// TIA Portal project "Tes simulation extract_V15.1" (V15.1) (continued)
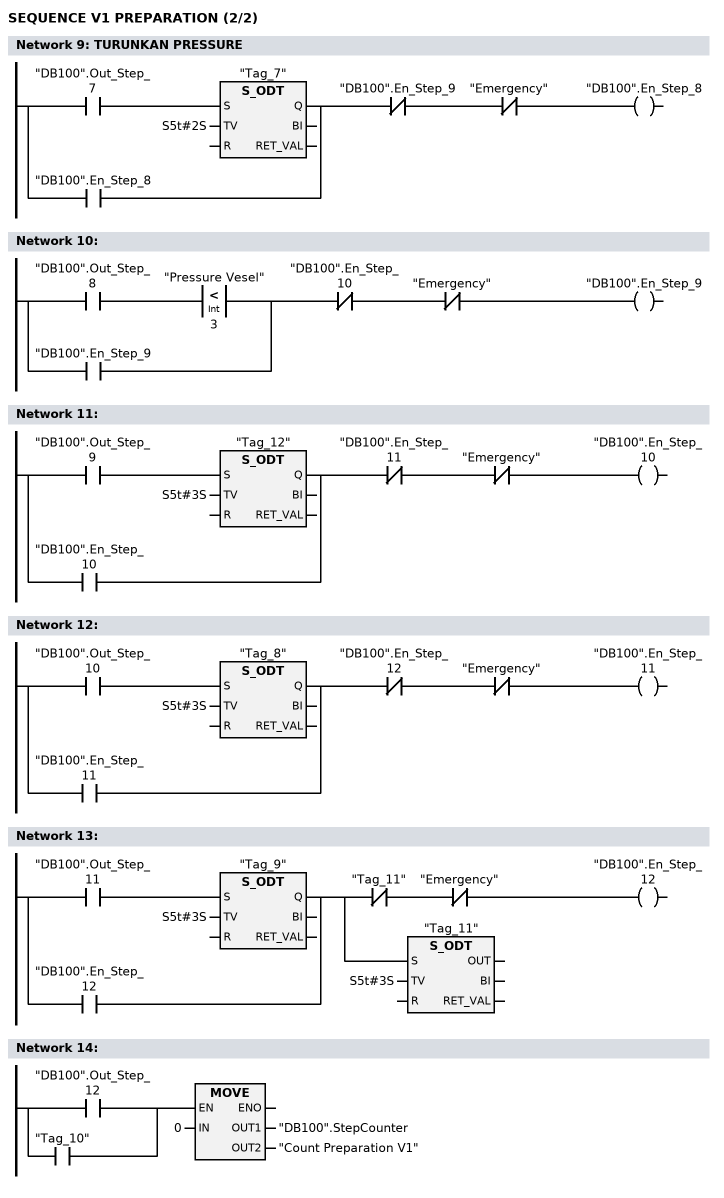
   RUNG wire#powerrail
      Contact( "DB100".Out_Step_7 )
      S_ODT(T_NO := "Tag_7", TV := S5t#2S, R :=, BI =>, RET_VAL =>)
      wire#w1
      I_Contact( "DB100".En_Step_9 )
      I_Contact( "Emergency" )
      Coil( "DB100".En_Step_8 )
   END_RUNG
   RUNG wire#powerrail
      Contact( "DB100".En_Step_8 )
   END_RUNG wire#w1
   // the same network as SCL:
   #_s5time1 := S_ODT(T_NO := "Tag_7", S := "DB100".Out_Step_7, TV := S5t#2S, Q => #_w1);
   "DB100".En_Step_8 := (#_w1 OR "DB100".En_Step_8) AND NOT "DB100".En_Step_9 AND NOT "Emergency";
END_REGION

REGION Network 10
   RUNG wire#powerrail
      Contact( "DB100".Out_Step_8 )
      { S7_Templates := "SrcType := Int" } LT_Contact(in1 := "Pressure Vesel", in2 := 3)
      wire#w1
      I_Contact( "DB100".En_Step_10 )
      I_Contact( "Emergency" )
      Coil( "DB100".En_Step_9 )
   END_RUNG
   RUNG wire#powerrail
      Contact( "DB100".En_Step_9 )
   END_RUNG wire#w1
   // the same network as SCL:
   "DB100".En_Step_9 := (("DB100".Out_Step_8 AND ("Pressure Vesel" < 3)) OR "DB100".En_Step_9) AND NOT "DB100".En_Step_10 AND NOT "Emergency";
END_REGION

REGION Network 11
   RUNG wire#powerrail
      Contact( "DB100".Out_Step_9 )
      S_ODT(T_NO := "Tag_12", TV := S5t#3S, R :=, BI =>, RET_VAL =>)
      wire#w1
      I_Contact( "DB100".En_Step_11 )
      I_Contact( "Emergency" )
      Coil( "DB100".En_Step_10 )
   END_RUNG
   RUNG wire#powerrail
      Contact( "DB100".En_Step_10 )
   END_RUNG wire#w1
   // the same network as SCL:
   #_s5time1 := S_ODT(T_NO := "Tag_12", S := "DB100".Out_Step_9, TV := S5t#3S, Q => #_w1);
   "DB100".En_Step_10 := (#_w1 OR "DB100".En_Step_10) AND NOT "DB100".En_Step_11 AND NOT "Emergency";
END_REGION

REGION Network 12
   RUNG wire#powerrail
      Contact( "DB100".Out_Step_10 )
      S_ODT(T_NO := "Tag_8", TV := S5t#3S, R :=, BI =>, RET_VAL =>)
      wire#w1
      I_Contact( "DB100".En_Step_12 )
      I_Contact( "Emergency" )
      Coil( "DB100".En_Step_11 )
   END_RUNG
   RUNG wire#powerrail
      Contact( "DB100".En_Step_11 )
   END_RUNG wire#w1
   // the same network as SCL:
   #_s5time1 := S_ODT(T_NO := "Tag_8", S := "DB100".Out_Step_10, TV := S5t#3S, Q => #_w1);
   "DB100".En_Step_11 := (#_w1 OR "DB100".En_Step_11) AND NOT "DB100".En_Step_12 AND NOT "Emergency";
END_REGION

REGION Network 13
   RUNG wire#powerrail
      Contact( "DB100".Out_Step_11 )
      S_ODT(T_NO := "Tag_9", TV := S5t#3S, R :=, BI =>, RET_VAL =>)
      wire#w1
      I_Contact( "Tag_11" )
      I_Contact( "Emergency" )
      Coil( "DB100".En_Step_12 )
   END_RUNG
   RUNG wire#powerrail
      Contact( "DB100".En_Step_12 )
   END_RUNG wire#w1
   RUNG wire#w1
      S_ODT(T_NO := "Tag_11", TV := S5t#3S, R :=, BI =>, RET_VAL =>)
   END_RUNG
   // the same network as SCL:
   #_s5time1 := S_ODT(T_NO := "Tag_9", S := "DB100".Out_Step_11, TV := S5t#3S, Q => #_w1);
   #_w2 := #_w1 OR "DB100".En_Step_12;
   "DB100".En_Step_12 := #_w2 AND NOT "Tag_11" AND NOT "Emergency";
   #_s5time2 := S_ODT(T_NO := "Tag_11", S := #_w2, TV := S5t#3S);
END_REGION

REGION Network 14
   RUNG wire#powerrail
      Contact( "DB100".Out_Step_12 )
      wire#w1
      Move(in := 0, out1 => "DB100".StepCounter, out2 => "Count Preparation V1")
   END_RUNG
   RUNG wire#powerrail
      Contact( "Tag_10" )
   END_RUNG wire#w1
   // the same network as SCL:
   IF "DB100".Out_Step_12 OR "Tag_10" THEN
       "DB100".StepCounter := 0;
       "Count Preparation V1" := 0;
   END_IF;
END_REGION
END_FUNCTION

FUNCTION "VESSEL 1 PREPARATION" : Void   // FC2, LAD
{ S7_Optimized_Access := 'TRUE' }
VERSION : 0.1
   VAR_TEMP   // added for the SCL form of the ladder/FBD networks
      _w1 : Bool;
      _w2 : Bool;
      _w3 : Bool;
      _w4 : Bool;
   END_VAR
BEGIN

REGION Network 1: NAIKAN PRESSURE STEAM
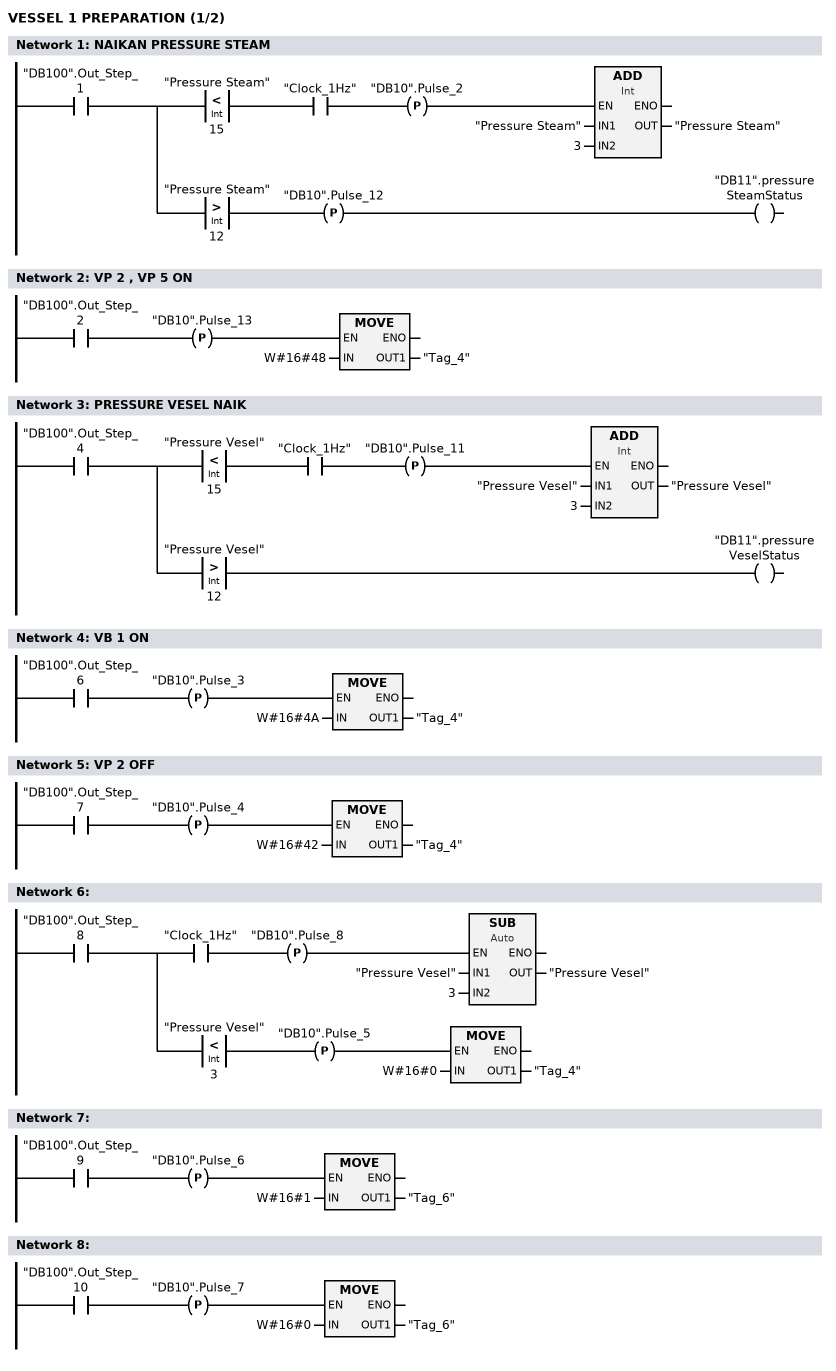
   RUNG wire#powerrail
      Contact( "DB100".Out_Step_1 )
      wire#w1
      { S7_Templates := "SrcType := Int" } LT_Contact(in1 := "Pressure Steam", in2 := 15)
      Contact( "Clock_1Hz" )
      P_Trig( "DB10".Pulse_2 )
      { S7_Templates := "SrcType := Int" } Add(in1 := "Pressure Steam", in2 := 3, out => "Pressure Steam")
   END_RUNG
   RUNG wire#w1
      { S7_Templates := "SrcType := Int" } GT_Contact(in1 := "Pressure Steam", in2 := 12)
      P_Trig( "DB10".Pulse_12 )
      Coil( "DB11".pressureSteamStatus )
   END_RUNG
   // the same network as SCL:
   #_w1 := "DB100".Out_Step_1 AND ("Pressure Steam" < 15) AND "Clock_1Hz";
   #_w2 := #_w1 AND NOT "DB10".Pulse_2;   // rising edge
   "DB10".Pulse_2 := #_w1;
   IF #_w2 THEN "Pressure Steam" := "Pressure Steam" + 3; END_IF;
   #_w3 := "DB100".Out_Step_1 AND ("Pressure Steam" > 12);
   #_w4 := #_w3 AND NOT "DB10".Pulse_12;   // rising edge
   "DB10".Pulse_12 := #_w3;
   "DB11".pressureSteamStatus := #_w4;
END_REGION

REGION Network 2: VP 2 , VP 5 ON
   RUNG wire#powerrail
      Contact( "DB100".Out_Step_2 )
      P_Trig( "DB10".Pulse_13 )
      Move(in := W#16#48, out1 => "Tag_4")
   END_RUNG
   // the same network as SCL:
   #_w1 := "DB100".Out_Step_2 AND NOT "DB10".Pulse_13;   // rising edge
   "DB10".Pulse_13 := "DB100".Out_Step_2;
   IF #_w1 THEN "Tag_4" := W#16#48; END_IF;
END_REGION

REGION Network 3: PRESSURE VESEL NAIK
   RUNG wire#powerrail
      Contact( "DB100".Out_Step_4 )
      wire#w1
      { S7_Templates := "SrcType := Int" } LT_Contact(in1 := "Pressure Vesel", in2 := 15)
      Contact( "Clock_1Hz" )
      P_Trig( "DB10".Pulse_11 )
      { S7_Templates := "SrcType := Int" } Add(in1 := "Pressure Vesel", in2 := 3, out => "Pressure Vesel")
   END_RUNG
   RUNG wire#w1
      { S7_Templates := "SrcType := Int" } GT_Contact(in1 := "Pressure Vesel", in2 := 12)
      Coil( "DB11".pressureVeselStatus )
   END_RUNG
   // the same network as SCL:
   #_w1 := "DB100".Out_Step_4 AND ("Pressure Vesel" < 15) AND "Clock_1Hz";
   #_w2 := #_w1 AND NOT "DB10".Pulse_11;   // rising edge
   "DB10".Pulse_11 := #_w1;
   IF #_w2 THEN "Pressure Vesel" := "Pressure Vesel" + 3; END_IF;
   "DB11".pressureVeselStatus := "DB100".Out_Step_4 AND ("Pressure Vesel" > 12);
END_REGION

REGION Network 4: VB 1 ON
   RUNG wire#powerrail
      Contact( "DB100".Out_Step_6 )
      P_Trig( "DB10".Pulse_3 )
      Move(in := W#16#4A, out1 => "Tag_4")
   END_RUNG
   // the same network as SCL:
   #_w1 := "DB100".Out_Step_6 AND NOT "DB10".Pulse_3;   // rising edge
   "DB10".Pulse_3 := "DB100".Out_Step_6;
   IF #_w1 THEN "Tag_4" := W#16#4A; END_IF;
END_REGION

REGION Network 5: VP 2 OFF
   RUNG wire#powerrail
      Contact( "DB100".Out_Step_7 )
      P_Trig( "DB10".Pulse_4 )
      Move(in := W#16#42, out1 => "Tag_4")
   END_RUNG
   // the same network as SCL:
   #_w1 := "DB100".Out_Step_7 AND NOT "DB10".Pulse_4;   // rising edge
   "DB10".Pulse_4 := "DB100".Out_Step_7;
   IF #_w1 THEN "Tag_4" := W#16#42; END_IF;
END_REGION

REGION Network 6
   RUNG wire#powerrail
      Contact( "DB100".Out_Step_8 )
      wire#w1
      Contact( "Clock_1Hz" )
      P_Trig( "DB10".Pulse_8 )
      Sub(in1 := "Pressure Vesel", in2 := 3, out => "Pressure Vesel")
   END_RUNG
   RUNG wire#w1
      { S7_Templates := "SrcType := Int" } LT_Contact(in1 := "Pressure Vesel", in2 := 3)
      P_Trig( "DB10".Pulse_5 )
      Move(in := W#16#0, out1 => "Tag_4")
   END_RUNG
   // the same network as SCL:
   #_w1 := "DB100".Out_Step_8 AND "Clock_1Hz";
   #_w2 := #_w1 AND NOT "DB10".Pulse_8;   // rising edge
   "DB10".Pulse_8 := #_w1;
   IF #_w2 THEN "Pressure Vesel" := "Pressure Vesel" - 3; END_IF;
   #_w3 := "DB100".Out_Step_8 AND ("Pressure Vesel" < 3);
   #_w4 := #_w3 AND NOT "DB10".Pulse_5;   // rising edge
   "DB10".Pulse_5 := #_w3;
   IF #_w4 THEN "Tag_4" := W#16#0; END_IF;
END_REGION

REGION Network 7
   RUNG wire#powerrail
      Contact( "DB100".Out_Step_9 )
      P_Trig( "DB10".Pulse_6 )
      Move(in := W#16#1, out1 => "Tag_6")
   END_RUNG
   // the same network as SCL:
   #_w1 := "DB100".Out_Step_9 AND NOT "DB10".Pulse_6;   // rising edge
   "DB10".Pulse_6 := "DB100".Out_Step_9;
   IF #_w1 THEN "Tag_6" := W#16#1; END_IF;
END_REGION

REGION Network 8
   RUNG wire#powerrail
      Contact( "DB100".Out_Step_10 )
      P_Trig( "DB10".Pulse_7 )
      Move(in := W#16#0, out1 => "Tag_6")
   END_RUNG
   // the same network as SCL:
   #_w1 := "DB100".Out_Step_10 AND NOT "DB10".Pulse_7;   // rising edge
   "DB10".Pulse_7 := "DB100".Out_Step_10;
   IF #_w1 THEN "Tag_6" := W#16#0; END_IF;
END_REGION

REGION Network 9
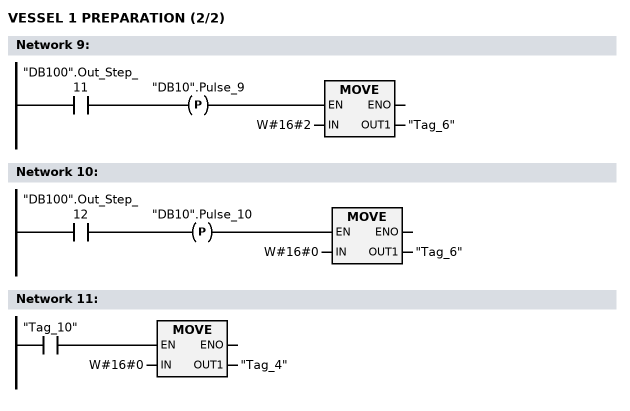
   RUNG wire#powerrail
      Contact( "DB100".Out_Step_11 )
      P_Trig( "DB10".Pulse_9 )
      Move(in := W#16#2, out1 => "Tag_6")
   END_RUNG
   // the same network as SCL:
   #_w1 := "DB100".Out_Step_11 AND NOT "DB10".Pulse_9;   // rising edge
   "DB10".Pulse_9 := "DB100".Out_Step_11;
   IF #_w1 THEN "Tag_6" := W#16#2; END_IF;
END_REGION

REGION Network 10
   RUNG wire#powerrail
      Contact( "DB100".Out_Step_12 )
      P_Trig( "DB10".Pulse_10 )
      Move(in := W#16#0, out1 => "Tag_6")
   END_RUNG
   // the same network as SCL:
   #_w1 := "DB100".Out_Step_12 AND NOT "DB10".Pulse_10;   // rising edge
   "DB10".Pulse_10 := "DB100".Out_Step_12;
   IF #_w1 THEN "Tag_6" := W#16#0; END_IF;
END_REGION

REGION Network 11
   RUNG wire#powerrail
      Contact( "Tag_10" )
      Move(in := W#16#0, out1 => "Tag_4")
   END_RUNG
   // the same network as SCL:
   IF "Tag_10" THEN "Tag_4" := W#16#0; END_IF;
END_REGION
END_FUNCTION

FUNCTION "ISI VESEL" : Void   // FC3, LAD
{ S7_Optimized_Access := 'TRUE' }
VERSION : 0.1
   VAR_TEMP   // added for the SCL form of the ladder/FBD networks
      _w1 : Bool;
      _w2 : Bool;
      _s5time1 : S5Time;
   END_VAR
BEGIN

REGION Network 1: ISI VESEL 1
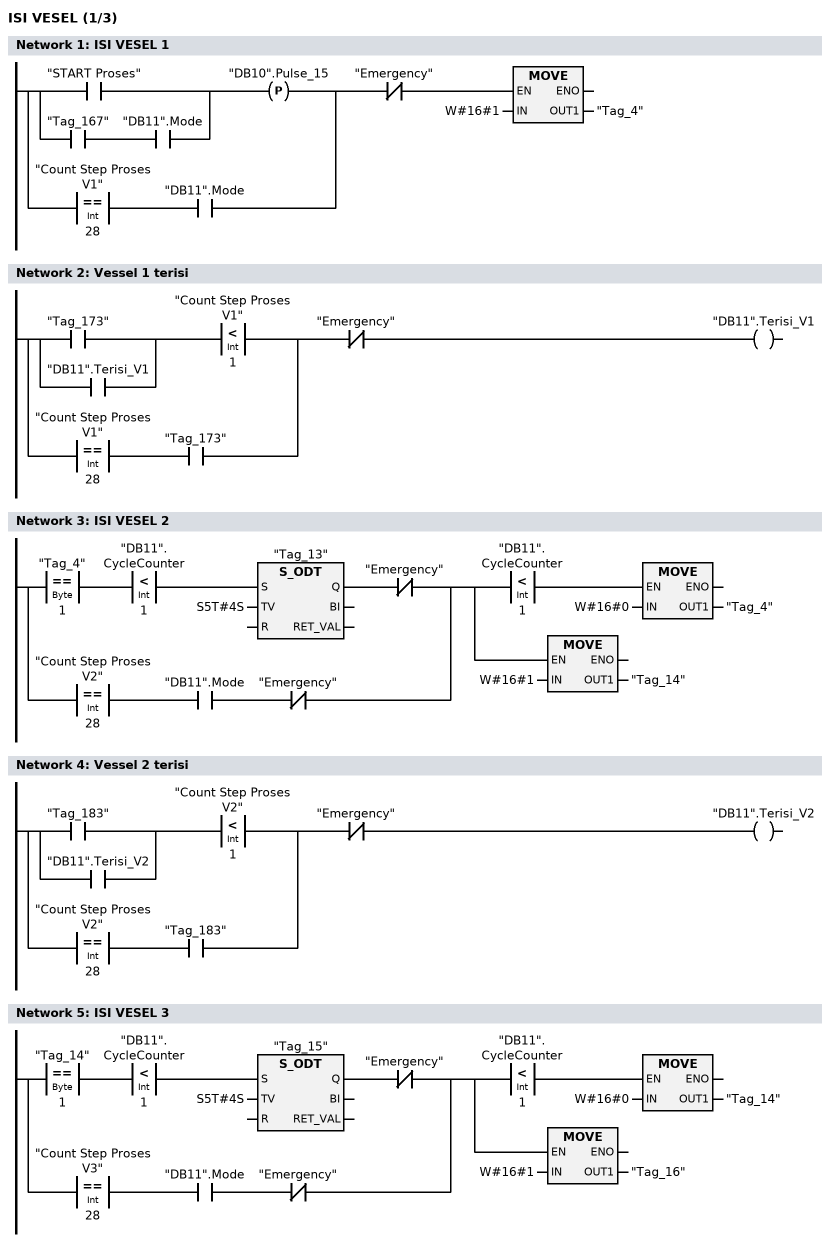
   RUNG wire#powerrail
      Contact( "START Proses" )
      wire#w1
      P_Trig( "DB10".Pulse_15 )
      wire#w2
      I_Contact( "Emergency" )
      Move(in := W#16#1, out1 => "Tag_4")
   END_RUNG
   RUNG wire#powerrail
      Contact( "Tag_167" )
      Contact( "DB11".Mode )
   END_RUNG wire#w1
   RUNG wire#powerrail
      { S7_Templates := "SrcType := Int" } EQ_Contact(in1 := "Count Step Proses V1", in2 := 28)
      Contact( "DB11".Mode )
   END_RUNG wire#w2
   // the same network as SCL:
   #_w1 := "START Proses" OR ("Tag_167" AND "DB11".Mode);
   #_w2 := #_w1 AND NOT "DB10".Pulse_15;   // rising edge
   "DB10".Pulse_15 := #_w1;
   IF (#_w2 OR (("Count Step Proses V1" = 28) AND "DB11".Mode)) AND NOT "Emergency" THEN
       "Tag_4" := W#16#1;
   END_IF;
END_REGION

REGION Network 2: Vessel 1 terisi
   RUNG wire#powerrail
      Contact( "Tag_173" )
      wire#w1
      { S7_Templates := "SrcType := Int" } LT_Contact(in1 := "Count Step Proses V1", in2 := 1)
      wire#w2
      I_Contact( "Emergency" )
      Coil( "DB11".Terisi_V1 )
   END_RUNG
   RUNG wire#powerrail
      Contact( "DB11".Terisi_V1 )
   END_RUNG wire#w1
   RUNG wire#powerrail
      { S7_Templates := "SrcType := Int" } EQ_Contact(in1 := "Count Step Proses V1", in2 := 28)
      Contact( "Tag_173" )
   END_RUNG wire#w2
   // the same network as SCL:
   "DB11".Terisi_V1 := ((("Tag_173" OR "DB11".Terisi_V1) AND ("Count Step Proses V1" < 1)) OR (("Count Step Proses V1" = 28) AND "Tag_173")) AND NOT "Emergency";
END_REGION

REGION Network 3: ISI VESEL 2
   RUNG wire#powerrail
      { S7_Templates := "SrcType := Byte" } EQ_Contact(in1 := "Tag_4", in2 := 1)
      { S7_Templates := "SrcType := Int" } LT_Contact(in1 := "DB11".CycleCounter, in2 := 1)
      S_ODT(T_NO := "Tag_13", TV := S5T#4S, R :=, BI =>, RET_VAL =>)
      I_Contact( "Emergency" )
      wire#w1
      { S7_Templates := "SrcType := Int" } LT_Contact(in1 := "DB11".CycleCounter, in2 := 1)
      Move(in := W#16#0, out1 => "Tag_4")
   END_RUNG
   RUNG wire#powerrail
      { S7_Templates := "SrcType := Int" } EQ_Contact(in1 := "Count Step Proses V2", in2 := 28)
      Contact( "DB11".Mode )
      I_Contact( "Emergency" )
   END_RUNG wire#w1
   RUNG wire#w1
      Move(in := W#16#1, out1 => "Tag_14")
   END_RUNG
   // the same network as SCL:
   #_s5time1 := S_ODT(T_NO := "Tag_13",
                      S := ("Tag_4" = 1) AND ("DB11".CycleCounter < 1),
                      TV := S5T#4S,
                      Q => #_w1);
   #_w2 := (#_w1 AND NOT "Emergency") OR (("Count Step Proses V2" = 28) AND "DB11".Mode AND NOT "Emergency");
   IF #_w2 AND ("DB11".CycleCounter < 1) THEN "Tag_4" := W#16#0; END_IF;
   IF #_w2 THEN "Tag_14" := W#16#1; END_IF;
END_REGION

REGION Network 4: Vessel 2 terisi
   RUNG wire#powerrail
      Contact( "Tag_183" )
      wire#w1
      { S7_Templates := "SrcType := Int" } LT_Contact(in1 := "Count Step Proses V2", in2 := 1)
      wire#w2
      I_Contact( "Emergency" )
      Coil( "DB11".Terisi_V2 )
   END_RUNG
   RUNG wire#powerrail
      Contact( "DB11".Terisi_V2 )
   END_RUNG wire#w1
   RUNG wire#powerrail
      { S7_Templates := "SrcType := Int" } EQ_Contact(in1 := "Count Step Proses V2", in2 := 28)
      Contact( "Tag_183" )
   END_RUNG wire#w2
   // the same network as SCL:
   "DB11".Terisi_V2 := ((("Tag_183" OR "DB11".Terisi_V2) AND ("Count Step Proses V2" < 1)) OR (("Count Step Proses V2" = 28) AND "Tag_183")) AND NOT "Emergency";
END_REGION

REGION Network 5: ISI VESEL 3
   RUNG wire#powerrail
      { S7_Templates := "SrcType := Byte" } EQ_Contact(in1 := "Tag_14", in2 := 1)
      { S7_Templates := "SrcType := Int" } LT_Contact(in1 := "DB11".CycleCounter, in2 := 1)
      S_ODT(T_NO := "Tag_15", TV := S5T#4S, R :=, BI =>, RET_VAL =>)
      I_Contact( "Emergency" )
      wire#w1
      { S7_Templates := "SrcType := Int" } LT_Contact(in1 := "DB11".CycleCounter, in2 := 1)
      Move(in := W#16#0, out1 => "Tag_14")
   END_RUNG
   RUNG wire#powerrail
      { S7_Templates := "SrcType := Int" } EQ_Contact(in1 := "Count Step Proses V3", in2 := 28)
      Contact( "DB11".Mode )
      I_Contact( "Emergency" )
   END_RUNG wire#w1
   RUNG wire#w1
      Move(in := W#16#1, out1 => "Tag_16")
   END_RUNG
   // the same network as SCL:
   #_s5time1 := S_ODT(T_NO := "Tag_15",
                      S := ("Tag_14" = 1) AND ("DB11".CycleCounter < 1),
                      TV := S5T#4S,
                      Q => #_w1);
   #_w2 := (#_w1 AND NOT "Emergency") OR (("Count Step Proses V3" = 28) AND "DB11".Mode AND NOT "Emergency");
   IF #_w2 AND ("DB11".CycleCounter < 1) THEN "Tag_14" := W#16#0; END_IF;
   IF #_w2 THEN "Tag_16" := W#16#1; END_IF;
END_REGION

REGION Network 6: Vessel 3 terisi
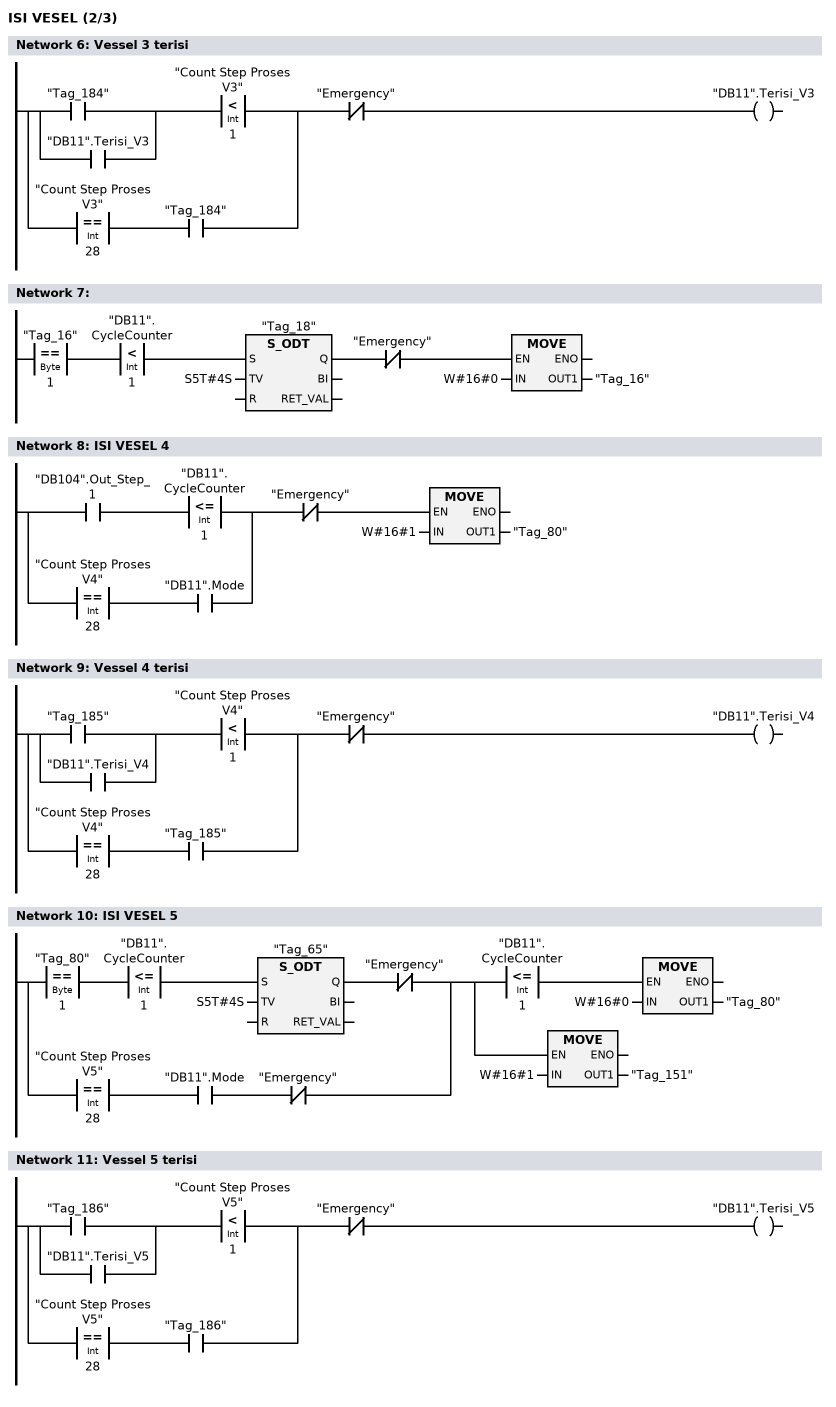
   RUNG wire#powerrail
      Contact( "Tag_184" )
      wire#w1
      { S7_Templates := "SrcType := Int" } LT_Contact(in1 := "Count Step Proses V3", in2 := 1)
      wire#w2
      I_Contact( "Emergency" )
      Coil( "DB11".Terisi_V3 )
   END_RUNG
   RUNG wire#powerrail
      Contact( "DB11".Terisi_V3 )
   END_RUNG wire#w1
   RUNG wire#powerrail
      { S7_Templates := "SrcType := Int" } EQ_Contact(in1 := "Count Step Proses V3", in2 := 28)
      Contact( "Tag_184" )
   END_RUNG wire#w2
   // the same network as SCL:
   "DB11".Terisi_V3 := ((("Tag_184" OR "DB11".Terisi_V3) AND ("Count Step Proses V3" < 1)) OR (("Count Step Proses V3" = 28) AND "Tag_184")) AND NOT "Emergency";
END_REGION

REGION Network 7
   RUNG wire#powerrail
      { S7_Templates := "SrcType := Byte" } EQ_Contact(in1 := "Tag_16", in2 := 1)
      { S7_Templates := "SrcType := Int" } LT_Contact(in1 := "DB11".CycleCounter, in2 := 1)
      S_ODT(T_NO := "Tag_18", TV := S5T#4S, R :=, BI =>, RET_VAL =>)
      I_Contact( "Emergency" )
      Move(in := W#16#0, out1 => "Tag_16")
   END_RUNG
   // the same network as SCL:
   #_s5time1 := S_ODT(T_NO := "Tag_18",
                      S := ("Tag_16" = 1) AND ("DB11".CycleCounter < 1),
                      TV := S5T#4S,
                      Q => #_w1);
   IF #_w1 AND NOT "Emergency" THEN "Tag_16" := W#16#0; END_IF;
END_REGION

REGION Network 8: ISI VESEL 4
   RUNG wire#powerrail
      Contact( "DB104".Out_Step_1 )
      { S7_Templates := "SrcType := Int" } LE_Contact(in1 := "DB11".CycleCounter, in2 := 1)
      wire#w1
      I_Contact( "Emergency" )
      Move(in := W#16#1, out1 => "Tag_80")
   END_RUNG
   RUNG wire#powerrail
      { S7_Templates := "SrcType := Int" } EQ_Contact(in1 := "Count Step Proses V4", in2 := 28)
      Contact( "DB11".Mode )
   END_RUNG wire#w1
   // the same network as SCL:
   IF (("DB104".Out_Step_1 AND ("DB11".CycleCounter <= 1)) OR (("Count Step Proses V4" = 28) AND "DB11".Mode)) AND NOT "Emergency" THEN
       "Tag_80" := W#16#1;
   END_IF;
END_REGION

REGION Network 9: Vessel 4 terisi
   RUNG wire#powerrail
      Contact( "Tag_185" )
      wire#w1
      { S7_Templates := "SrcType := Int" } LT_Contact(in1 := "Count Step Proses V4", in2 := 1)
      wire#w2
      I_Contact( "Emergency" )
      Coil( "DB11".Terisi_V4 )
   END_RUNG
   RUNG wire#powerrail
      Contact( "DB11".Terisi_V4 )
   END_RUNG wire#w1
   RUNG wire#powerrail
      { S7_Templates := "SrcType := Int" } EQ_Contact(in1 := "Count Step Proses V4", in2 := 28)
      Contact( "Tag_185" )
   END_RUNG wire#w2
   // the same network as SCL:
   "DB11".Terisi_V4 := ((("Tag_185" OR "DB11".Terisi_V4) AND ("Count Step Proses V4" < 1)) OR (("Count Step Proses V4" = 28) AND "Tag_185")) AND NOT "Emergency";
END_REGION

REGION Network 10: ISI VESEL 5
   RUNG wire#powerrail
      { S7_Templates := "SrcType := Byte" } EQ_Contact(in1 := "Tag_80", in2 := 1)
      { S7_Templates := "SrcType := Int" } LE_Contact(in1 := "DB11".CycleCounter, in2 := 1)
      S_ODT(T_NO := "Tag_65", TV := S5T#4S, R :=, BI =>, RET_VAL =>)
      I_Contact( "Emergency" )
      wire#w1
      { S7_Templates := "SrcType := Int" } LE_Contact(in1 := "DB11".CycleCounter, in2 := 1)
      Move(in := W#16#0, out1 => "Tag_80")
   END_RUNG
   RUNG wire#powerrail
      { S7_Templates := "SrcType := Int" } EQ_Contact(in1 := "Count Step Proses V5", in2 := 28)
      Contact( "DB11".Mode )
      I_Contact( "Emergency" )
   END_RUNG wire#w1
   RUNG wire#w1
      Move(in := W#16#1, out1 => "Tag_151")
   END_RUNG
   // the same network as SCL:
   #_s5time1 := S_ODT(T_NO := "Tag_65",
                      S := ("Tag_80" = 1) AND ("DB11".CycleCounter <= 1),
                      TV := S5T#4S,
                      Q => #_w1);
   #_w2 := (#_w1 AND NOT "Emergency") OR (("Count Step Proses V5" = 28) AND "DB11".Mode AND NOT "Emergency");
   IF #_w2 AND ("DB11".CycleCounter <= 1) THEN "Tag_80" := W#16#0; END_IF;
   IF #_w2 THEN "Tag_151" := W#16#1; END_IF;
END_REGION

REGION Network 11: Vessel 5 terisi
   RUNG wire#powerrail
      Contact( "Tag_186" )
      wire#w1
      { S7_Templates := "SrcType := Int" } LT_Contact(in1 := "Count Step Proses V5", in2 := 1)
      wire#w2
      I_Contact( "Emergency" )
      Coil( "DB11".Terisi_V5 )
   END_RUNG
   RUNG wire#powerrail
      Contact( "DB11".Terisi_V5 )
   END_RUNG wire#w1
   RUNG wire#powerrail
      { S7_Templates := "SrcType := Int" } EQ_Contact(in1 := "Count Step Proses V5", in2 := 28)
      Contact( "Tag_186" )
   END_RUNG wire#w2
   // the same network as SCL:
   "DB11".Terisi_V5 := ((("Tag_186" OR "DB11".Terisi_V5) AND ("Count Step Proses V5" < 1)) OR (("Count Step Proses V5" = 28) AND "Tag_186")) AND NOT "Emergency";
END_REGION

REGION Network 12: ISI VESEL 6
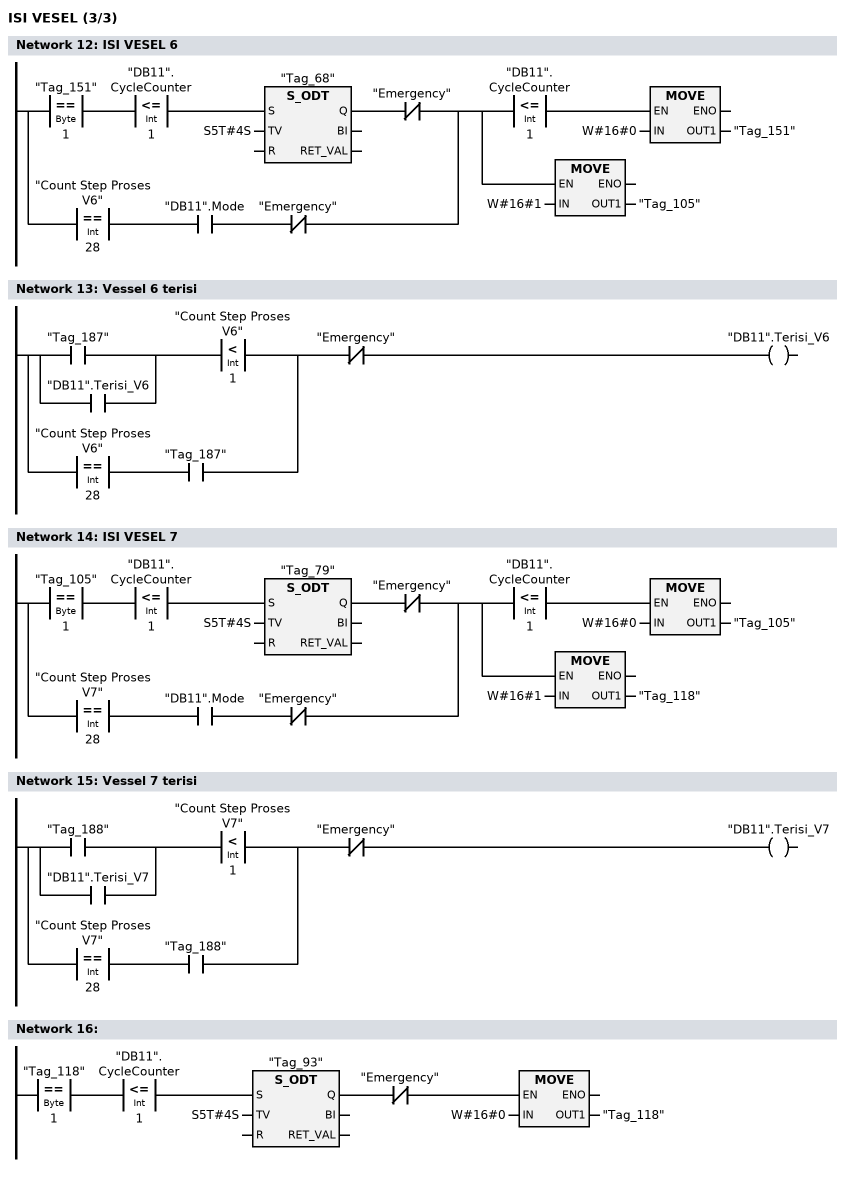
   RUNG wire#powerrail
      { S7_Templates := "SrcType := Byte" } EQ_Contact(in1 := "Tag_151", in2 := 1)
      { S7_Templates := "SrcType := Int" } LE_Contact(in1 := "DB11".CycleCounter, in2 := 1)
      S_ODT(T_NO := "Tag_68", TV := S5T#4S, R :=, BI =>, RET_VAL =>)
      I_Contact( "Emergency" )
      wire#w1
      { S7_Templates := "SrcType := Int" } LE_Contact(in1 := "DB11".CycleCounter, in2 := 1)
      Move(in := W#16#0, out1 => "Tag_151")
   END_RUNG
   RUNG wire#powerrail
      { S7_Templates := "SrcType := Int" } EQ_Contact(in1 := "Count Step Proses V6", in2 := 28)
      Contact( "DB11".Mode )
      I_Contact( "Emergency" )
   END_RUNG wire#w1
   RUNG wire#w1
      Move(in := W#16#1, out1 => "Tag_105")
   END_RUNG
   // the same network as SCL:
   #_s5time1 := S_ODT(T_NO := "Tag_68",
                      S := ("Tag_151" = 1) AND ("DB11".CycleCounter <= 1),
                      TV := S5T#4S,
                      Q => #_w1);
   #_w2 := (#_w1 AND NOT "Emergency") OR (("Count Step Proses V6" = 28) AND "DB11".Mode AND NOT "Emergency");
   IF #_w2 AND ("DB11".CycleCounter <= 1) THEN "Tag_151" := W#16#0; END_IF;
   IF #_w2 THEN "Tag_105" := W#16#1; END_IF;
END_REGION

REGION Network 13: Vessel 6 terisi
   RUNG wire#powerrail
      Contact( "Tag_187" )
      wire#w1
      { S7_Templates := "SrcType := Int" } LT_Contact(in1 := "Count Step Proses V6", in2 := 1)
      wire#w2
      I_Contact( "Emergency" )
      Coil( "DB11".Terisi_V6 )
   END_RUNG
   RUNG wire#powerrail
      Contact( "DB11".Terisi_V6 )
   END_RUNG wire#w1
   RUNG wire#powerrail
      { S7_Templates := "SrcType := Int" } EQ_Contact(in1 := "Count Step Proses V6", in2 := 28)
      Contact( "Tag_187" )
   END_RUNG wire#w2
   // the same network as SCL:
   "DB11".Terisi_V6 := ((("Tag_187" OR "DB11".Terisi_V6) AND ("Count Step Proses V6" < 1)) OR (("Count Step Proses V6" = 28) AND "Tag_187")) AND NOT "Emergency";
END_REGION

REGION Network 14: ISI VESEL 7
   RUNG wire#powerrail
      { S7_Templates := "SrcType := Byte" } EQ_Contact(in1 := "Tag_105", in2 := 1)
      { S7_Templates := "SrcType := Int" } LE_Contact(in1 := "DB11".CycleCounter, in2 := 1)
      S_ODT(T_NO := "Tag_79", TV := S5T#4S, R :=, BI =>, RET_VAL =>)
      I_Contact( "Emergency" )
      wire#w1
      { S7_Templates := "SrcType := Int" } LE_Contact(in1 := "DB11".CycleCounter, in2 := 1)
      Move(in := W#16#0, out1 => "Tag_105")
   END_RUNG
   RUNG wire#powerrail
      { S7_Templates := "SrcType := Int" } EQ_Contact(in1 := "Count Step Proses V7", in2 := 28)
      Contact( "DB11".Mode )
      I_Contact( "Emergency" )
   END_RUNG wire#w1
   RUNG wire#w1
      Move(in := W#16#1, out1 => "Tag_118")
   END_RUNG
   // the same network as SCL:
   #_s5time1 := S_ODT(T_NO := "Tag_79",
                      S := ("Tag_105" = 1) AND ("DB11".CycleCounter <= 1),
                      TV := S5T#4S,
                      Q => #_w1);
   #_w2 := (#_w1 AND NOT "Emergency") OR (("Count Step Proses V7" = 28) AND "DB11".Mode AND NOT "Emergency");
   IF #_w2 AND ("DB11".CycleCounter <= 1) THEN "Tag_105" := W#16#0; END_IF;
   IF #_w2 THEN "Tag_118" := W#16#1; END_IF;
END_REGION

REGION Network 15: Vessel 7 terisi
   RUNG wire#powerrail
      Contact( "Tag_188" )
      wire#w1
      { S7_Templates := "SrcType := Int" } LT_Contact(in1 := "Count Step Proses V7", in2 := 1)
      wire#w2
      I_Contact( "Emergency" )
      Coil( "DB11".Terisi_V7 )
   END_RUNG
   RUNG wire#powerrail
      Contact( "DB11".Terisi_V7 )
   END_RUNG wire#w1
   RUNG wire#powerrail
      { S7_Templates := "SrcType := Int" } EQ_Contact(in1 := "Count Step Proses V7", in2 := 28)
      Contact( "Tag_188" )
   END_RUNG wire#w2
   // the same network as SCL:
   "DB11".Terisi_V7 := ((("Tag_188" OR "DB11".Terisi_V7) AND ("Count Step Proses V7" < 1)) OR (("Count Step Proses V7" = 28) AND "Tag_188")) AND NOT "Emergency";
END_REGION

REGION Network 16
   RUNG wire#powerrail
      { S7_Templates := "SrcType := Byte" } EQ_Contact(in1 := "Tag_118", in2 := 1)
      { S7_Templates := "SrcType := Int" } LE_Contact(in1 := "DB11".CycleCounter, in2 := 1)
      S_ODT(T_NO := "Tag_93", TV := S5T#4S, R :=, BI =>, RET_VAL =>)
      I_Contact( "Emergency" )
      Move(in := W#16#0, out1 => "Tag_118")
   END_RUNG
   // the same network as SCL:
   #_s5time1 := S_ODT(T_NO := "Tag_93",
                      S := ("Tag_118" = 1) AND ("DB11".CycleCounter <= 1),
                      TV := S5T#4S,
                      Q => #_w1);
   IF #_w1 AND NOT "Emergency" THEN "Tag_118" := W#16#0; END_IF;
END_REGION
END_FUNCTION

FUNCTION "SUPPLY" : Void   // FC4, LAD
{ S7_Optimized_Access := 'TRUE' }
VERSION : 0.1
   VAR_TEMP   // added for the SCL form of the ladder/FBD networks
      _w1 : Bool;
      _w2 : Bool;
      _w3 : Bool;
      _w4 : Bool;
   END_VAR
BEGIN

REGION Network 1: BUKA CV AIR 1
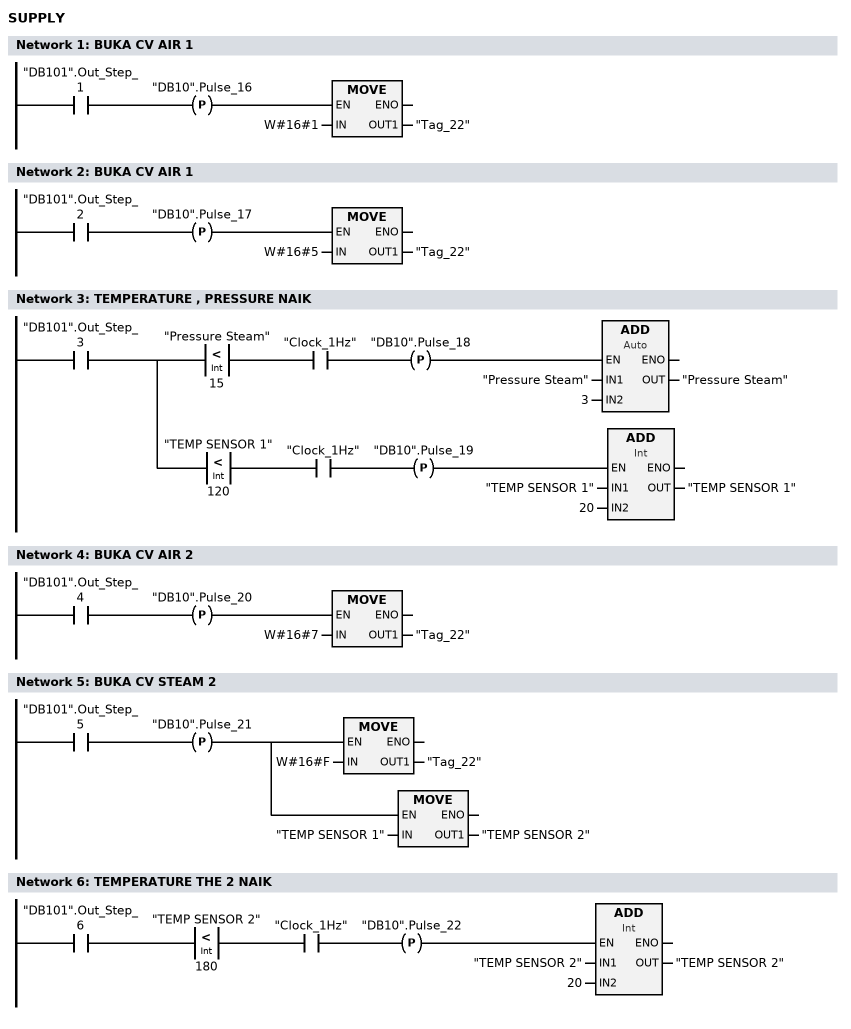
   RUNG wire#powerrail
      Contact( "DB101".Out_Step_1 )
      P_Trig( "DB10".Pulse_16 )
      Move(in := W#16#1, out1 => "Tag_22")
   END_RUNG
   // the same network as SCL:
   #_w1 := "DB101".Out_Step_1 AND NOT "DB10".Pulse_16;   // rising edge
   "DB10".Pulse_16 := "DB101".Out_Step_1;
   IF #_w1 THEN "Tag_22" := W#16#1; END_IF;
END_REGION

REGION Network 2: BUKA CV AIR 1
   RUNG wire#powerrail
      Contact( "DB101".Out_Step_2 )
      P_Trig( "DB10".Pulse_17 )
      Move(in := W#16#5, out1 => "Tag_22")
   END_RUNG
   // the same network as SCL:
   #_w1 := "DB101".Out_Step_2 AND NOT "DB10".Pulse_17;   // rising edge
   "DB10".Pulse_17 := "DB101".Out_Step_2;
   IF #_w1 THEN "Tag_22" := W#16#5; END_IF;
END_REGION

REGION Network 3: TEMPERATURE , PRESSURE NAIK
   RUNG wire#powerrail
      Contact( "DB101".Out_Step_3 )
      wire#w1
      { S7_Templates := "SrcType := Int" } LT_Contact(in1 := "Pressure Steam", in2 := 15)
      Contact( "Clock_1Hz" )
      P_Trig( "DB10".Pulse_18 )
      Add(in1 := "Pressure Steam", in2 := 3, out => "Pressure Steam")
   END_RUNG
   RUNG wire#w1
      { S7_Templates := "SrcType := Int" } LT_Contact(in1 := "TEMP SENSOR 1", in2 := 120)
      Contact( "Clock_1Hz" )
      P_Trig( "DB10".Pulse_19 )
      { S7_Templates := "SrcType := Int" } Add(in1 := "TEMP SENSOR 1", in2 := 20, out => "TEMP SENSOR 1")
   END_RUNG
   // the same network as SCL:
   #_w1 := "DB101".Out_Step_3 AND ("Pressure Steam" < 15) AND "Clock_1Hz";
   #_w2 := #_w1 AND NOT "DB10".Pulse_18;   // rising edge
   "DB10".Pulse_18 := #_w1;
   IF #_w2 THEN "Pressure Steam" := "Pressure Steam" + 3; END_IF;
   #_w3 := "DB101".Out_Step_3 AND ("TEMP SENSOR 1" < 120) AND "Clock_1Hz";
   #_w4 := #_w3 AND NOT "DB10".Pulse_19;   // rising edge
   "DB10".Pulse_19 := #_w3;
   IF #_w4 THEN "TEMP SENSOR 1" := "TEMP SENSOR 1" + 20; END_IF;
END_REGION

REGION Network 4: BUKA CV AIR 2
   RUNG wire#powerrail
      Contact( "DB101".Out_Step_4 )
      P_Trig( "DB10".Pulse_20 )
      Move(in := W#16#7, out1 => "Tag_22")
   END_RUNG
   // the same network as SCL:
   #_w1 := "DB101".Out_Step_4 AND NOT "DB10".Pulse_20;   // rising edge
   "DB10".Pulse_20 := "DB101".Out_Step_4;
   IF #_w1 THEN "Tag_22" := W#16#7; END_IF;
END_REGION

REGION Network 5: BUKA CV STEAM 2
   RUNG wire#powerrail
      Contact( "DB101".Out_Step_5 )
      P_Trig( "DB10".Pulse_21 )
      wire#w1
      Move(in := W#16#F, out1 => "Tag_22")
   END_RUNG
   RUNG wire#w1
      Move(in := "TEMP SENSOR 1", out1 => "TEMP SENSOR 2")
   END_RUNG
   // the same network as SCL:
   #_w1 := "DB101".Out_Step_5 AND NOT "DB10".Pulse_21;   // rising edge
   "DB10".Pulse_21 := "DB101".Out_Step_5;
   IF #_w1 THEN
       "Tag_22" := W#16#F;
       "TEMP SENSOR 2" := "TEMP SENSOR 1";
   END_IF;
END_REGION

REGION Network 6: TEMPERATURE THE 2 NAIK
   RUNG wire#powerrail
      Contact( "DB101".Out_Step_6 )
      { S7_Templates := "SrcType := Int" } LT_Contact(in1 := "TEMP SENSOR 2", in2 := 180)
      Contact( "Clock_1Hz" )
      P_Trig( "DB10".Pulse_22 )
      { S7_Templates := "SrcType := Int" } Add(in1 := "TEMP SENSOR 2", in2 := 20, out => "TEMP SENSOR 2")
   END_RUNG
   // the same network as SCL:
   #_w1 := "DB101".Out_Step_6 AND ("TEMP SENSOR 2" < 180) AND "Clock_1Hz";
   #_w2 := #_w1 AND NOT "DB10".Pulse_22;   // rising edge
   "DB10".Pulse_22 := #_w1;
   IF #_w2 THEN "TEMP SENSOR 2" := "TEMP SENSOR 2" + 20; END_IF;
END_REGION
END_FUNCTION

FUNCTION "SEQUENCE SUPPLY" : Void   // FC5, LAD
{ S7_Optimized_Access := 'TRUE' }
VERSION : 0.1
   VAR_TEMP   // added for the SCL form of the ladder/FBD networks
      _w1 : Bool;
      _s5time1 : S5Time;
   END_VAR
BEGIN

REGION Network 1: START SUPPLY
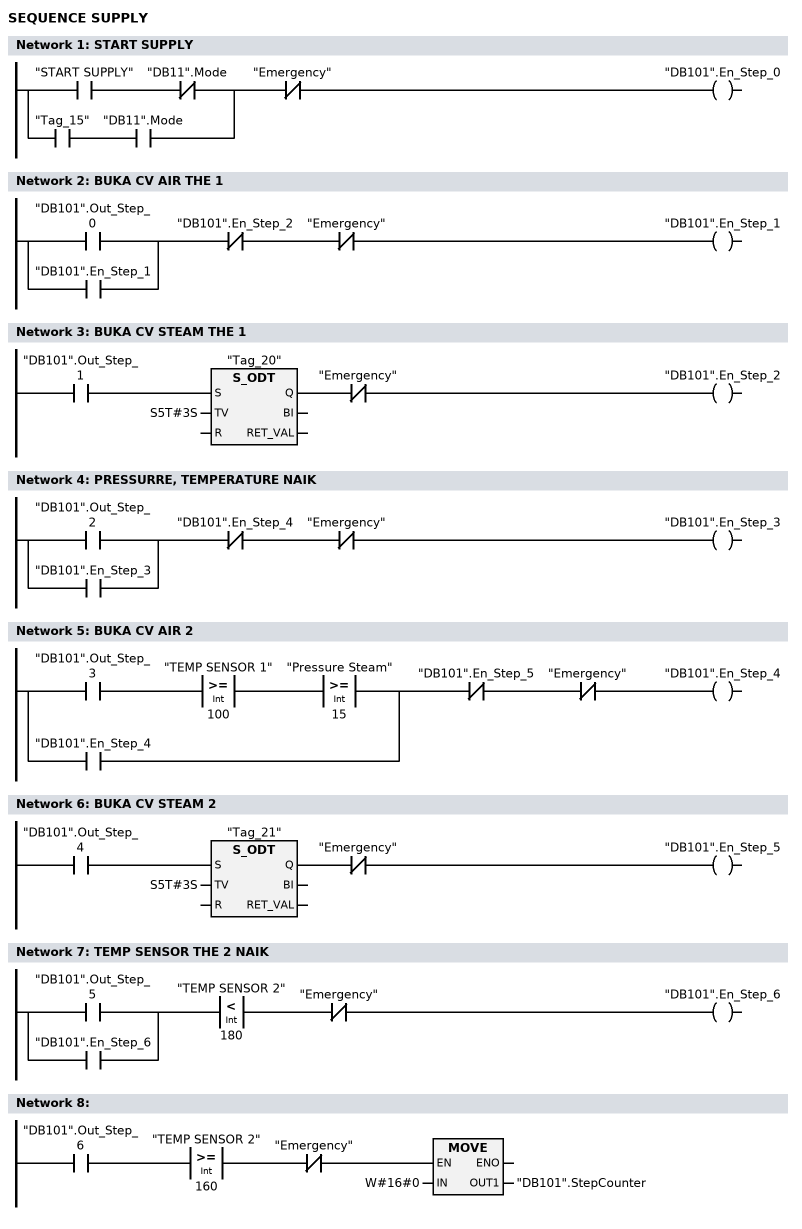
   RUNG wire#powerrail
      Contact( "START SUPPLY" )
      I_Contact( "DB11".Mode )
      wire#w1
      I_Contact( "Emergency" )
      Coil( "DB101".En_Step_0 )
   END_RUNG
   RUNG wire#powerrail
      Contact( "Tag_15" )
      Contact( "DB11".Mode )
   END_RUNG wire#w1
   // the same network as SCL:
   "DB101".En_Step_0 := (("START SUPPLY" AND NOT "DB11".Mode) OR ("Tag_15" AND "DB11".Mode)) AND NOT "Emergency";
END_REGION

REGION Network 2: BUKA CV AIR THE 1
   RUNG wire#powerrail
      Contact( "DB101".Out_Step_0 )
      wire#w1
      I_Contact( "DB101".En_Step_2 )
      I_Contact( "Emergency" )
      Coil( "DB101".En_Step_1 )
   END_RUNG
   RUNG wire#powerrail
      Contact( "DB101".En_Step_1 )
   END_RUNG wire#w1
   // the same network as SCL:
   "DB101".En_Step_1 := ("DB101".Out_Step_0 OR "DB101".En_Step_1) AND NOT "DB101".En_Step_2 AND NOT "Emergency";
END_REGION

REGION Network 3: BUKA CV STEAM THE 1
   RUNG wire#powerrail
      Contact( "DB101".Out_Step_1 )
      S_ODT(T_NO := "Tag_20", TV := S5T#3S, R :=, BI =>, RET_VAL =>)
      I_Contact( "Emergency" )
      Coil( "DB101".En_Step_2 )
   END_RUNG
   // the same network as SCL:
   #_s5time1 := S_ODT(T_NO := "Tag_20", S := "DB101".Out_Step_1, TV := S5T#3S, Q => #_w1);
   "DB101".En_Step_2 := #_w1 AND NOT "Emergency";
END_REGION

REGION Network 4: PRESSURRE, TEMPERATURE NAIK
   RUNG wire#powerrail
      Contact( "DB101".Out_Step_2 )
      wire#w1
      I_Contact( "DB101".En_Step_4 )
      I_Contact( "Emergency" )
      Coil( "DB101".En_Step_3 )
   END_RUNG
   RUNG wire#powerrail
      Contact( "DB101".En_Step_3 )
   END_RUNG wire#w1
   // the same network as SCL:
   "DB101".En_Step_3 := ("DB101".Out_Step_2 OR "DB101".En_Step_3) AND NOT "DB101".En_Step_4 AND NOT "Emergency";
END_REGION

REGION Network 5: BUKA CV AIR 2
   RUNG wire#powerrail
      Contact( "DB101".Out_Step_3 )
      { S7_Templates := "SrcType := Int" } GE_Contact(in1 := "TEMP SENSOR 1", in2 := 100)
      { S7_Templates := "SrcType := Int" } GE_Contact(in1 := "Pressure Steam", in2 := 15)
      wire#w1
      I_Contact( "DB101".En_Step_5 )
      I_Contact( "Emergency" )
      Coil( "DB101".En_Step_4 )
   END_RUNG
   RUNG wire#powerrail
      Contact( "DB101".En_Step_4 )
   END_RUNG wire#w1
   // the same network as SCL:
   "DB101".En_Step_4 := (("DB101".Out_Step_3 AND ("TEMP SENSOR 1" >= 100) AND ("Pressure Steam" >= 15)) OR "DB101".En_Step_4) AND NOT "DB101".En_Step_5 AND NOT "Emergency";
END_REGION

REGION Network 6: BUKA CV STEAM 2
   RUNG wire#powerrail
      Contact( "DB101".Out_Step_4 )
      S_ODT(T_NO := "Tag_21", TV := S5T#3S, R :=, BI =>, RET_VAL =>)
      I_Contact( "Emergency" )
      Coil( "DB101".En_Step_5 )
   END_RUNG
   // the same network as SCL:
   #_s5time1 := S_ODT(T_NO := "Tag_21", S := "DB101".Out_Step_4, TV := S5T#3S, Q => #_w1);
   "DB101".En_Step_5 := #_w1 AND NOT "Emergency";
END_REGION

REGION Network 7: TEMP SENSOR THE 2 NAIK
   RUNG wire#powerrail
      Contact( "DB101".Out_Step_5 )
      wire#w1
      { S7_Templates := "SrcType := Int" } LT_Contact(in1 := "TEMP SENSOR 2", in2 := 180)
      I_Contact( "Emergency" )
      Coil( "DB101".En_Step_6 )
   END_RUNG
   RUNG wire#powerrail
      Contact( "DB101".En_Step_6 )
   END_RUNG wire#w1
   // the same network as SCL:
   "DB101".En_Step_6 := ("DB101".Out_Step_5 OR "DB101".En_Step_6) AND ("TEMP SENSOR 2" < 180) AND NOT "Emergency";
END_REGION

REGION Network 8
   RUNG wire#powerrail
      Contact( "DB101".Out_Step_6 )
      { S7_Templates := "SrcType := Int" } GE_Contact(in1 := "TEMP SENSOR 2", in2 := 160)
      I_Contact( "Emergency" )
      Move(in := W#16#0, out1 => "DB101".StepCounter)
   END_RUNG
   // the same network as SCL:
   IF "DB101".Out_Step_6 AND ("TEMP SENSOR 2" >= 160) AND NOT "Emergency" THEN
       "DB101".StepCounter := W#16#0;
   END_IF;
END_REGION
END_FUNCTION

FUNCTION "VESSEL 1 PROSES" : Void   // FC6, LAD
{ S7_Optimized_Access := 'TRUE' }